// TIA Portal project "Semaforo Estruturado" (V16)

(* hardware
DEVICE "S7-1200 station_1"  S7-1200 Station
   slot 0: "Rack_0"  S7-1200 Rack  Rack  V1.0
   slot 1: "PLC_1"  CPU 1215C DC/DC/Rly  6ES7 215-1HG40-0XB0  V4.4
*)

// ===== PLC "PLC_1"  CPU 1215C DC/DC/Rly =====

VAR_GLOBAL   // PLC tag table "Default tag table"
   "Clock_Byte" AT %MB0 : Byte;
   "Clock_10Hz" AT %M0.0 : Bool;
   "Clock_5Hz" AT %M0.1 : Bool;
   "Clock_2.5Hz" AT %M0.2 : Bool;
   "Clock_2Hz" AT %M0.3 : Bool;
   "Clock_1.25Hz" AT %M0.4 : Bool;
   "Clock_1Hz" AT %M0.5 : Bool;
   "Clock_0.625Hz" AT %M0.6 : Bool;
   "Clock_0.5Hz" AT %M0.7 : Bool;
END_VAR

DATA_BLOCK "DB_Geral"   // DB1
{ S7_Optimized_Access := 'TRUE' }
VERSION : 0.1
   VAR
      Start : Bool;
      Stop : Bool;
      Reset : Bool;
      Estado : Bool;
      Time_of_Process : DInt;
      Time_PE_GroupA : Struct
         CutTimePE : DInt;
         TimePE : DInt := 20;
      END_STRUCT;
      Time_PE_GroupB : Struct
         CutTimePE : DInt;
         TimePE : DInt := 20;
      END_STRUCT;
      TimeOutCiclo : Struct
         "Estado 1" : DInt := 110;
         "Estado 2" : DInt := 120;
      END_STRUCT;
      ContadorGrupo : IEC_DCOUNTER;
   END_VAR
   VAR RETAIN
      PE : Struct
         GroupA : Bool;
         GroupB : Bool;
      END_STRUCT;
   END_VAR
   VAR
      Time_GroupA : Struct
         Red : Struct
            "begin" : DInt := 0;
            end : DInt := 40;
         END_STRUCT;
         Red_1 : Struct
            "begin" : DInt := 80;
            end : DInt := 110;
         END_STRUCT;
         Green : Struct
            "begin" : DInt := 40;
            end : DInt := 70;
         END_STRUCT;
         Yellow : Struct
            "begin" : DInt := 70;
            end : DInt := 80;
         END_STRUCT;
      END_STRUCT;
      Time_GroupB : Struct
         Red : Struct
            "begin" : DInt := 40;
            end : DInt := 110;
         END_STRUCT;
         Green : Struct
            "begin" : DInt := 0;
            end : DInt := 30;
         END_STRUCT;
         Yellow : Struct
            "begin" : DInt := 30;
            end : DInt := 40;
         END_STRUCT;
      END_STRUCT;
      Time_GroupC : Struct
         Red : Struct
            "begin" : DInt;
            end : DInt := 80;
         END_STRUCT;
         Green : Struct
            "begin" : DInt := 80;
            end : DInt := 100;
         END_STRUCT;
         Yellow : Struct
            "begin" : DInt := 100;
            end : DInt := 110;
         END_STRUCT;
      END_STRUCT;
   END_VAR
BEGIN
   ContadorGrupo.PV := 110;
END_DATA_BLOCK

DATA_BLOCK "DB_Input"   // DB2
{ S7_Optimized_Access := 'TRUE' }
VERSION : 0.1
   VAR
      Btn_PE_GroupA : Bool;
      Btn_PE_GroupB : Bool;
      Btn_Start : Bool;
      Btn_Stop : Bool;
      Btn_TestLamp : Bool;
      Btn_Reset : Bool;
   END_VAR
BEGIN
END_DATA_BLOCK

DATA_BLOCK "DB_Output"   // DB3
{ S7_Optimized_Access := 'TRUE' }
VERSION : 0.1
   VAR
      GroupA : Struct
         LampGreen : Bool;
         LampYell : Bool;
         LampRed : Bool;
      END_STRUCT;
      GroupB : Struct
         LampGreen : Bool;
         LampYell : Bool;
         LampRed : Bool;
      END_STRUCT;
      GroupC : Struct
         LampGreen : Bool;
         LampYell : Bool;
         LampRed : Bool;
      END_STRUCT;
      PE_GroupA : Struct
         LampGreen : Bool;
         LampRed : Bool;
      END_STRUCT;
      PE_GroupB : Struct
         LampGreen : Bool;
         LampRed : Bool;
      END_STRUCT;
   END_VAR
BEGIN
END_DATA_BLOCK

FUNCTION "FC_Geral" : Void   // FC1, LAD
{ S7_Optimized_Access := 'TRUE' }
VERSION : 0.1
   VAR_TEMP   // added for the SCL form of the ladder/FBD networks
      _w1 : Bool;
   END_VAR
BEGIN

REGION Network 1: Modo Start
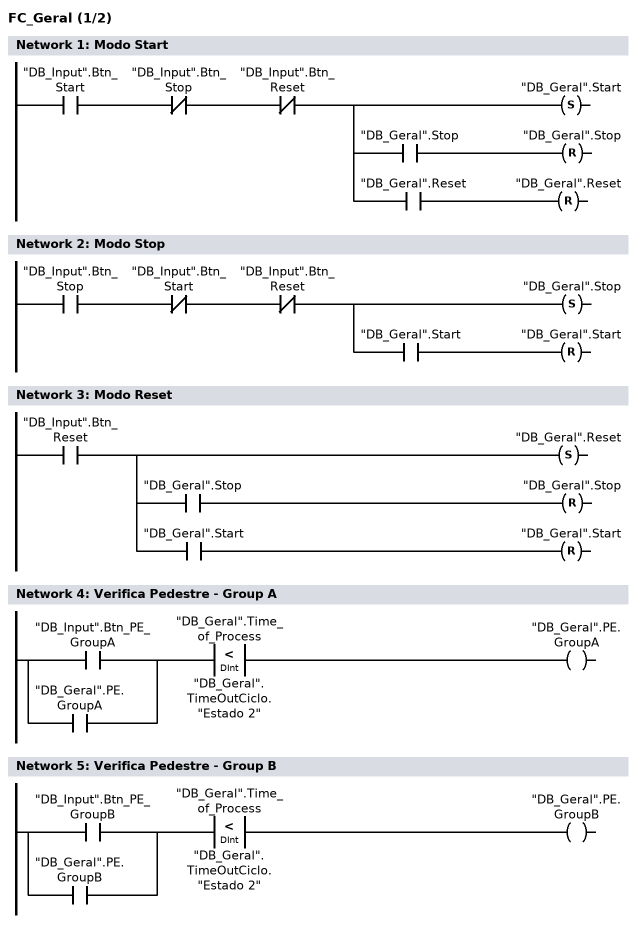
   RUNG wire#powerrail
      Contact( "DB_Input".Btn_Start )
      I_Contact( "DB_Input".Btn_Stop )
      I_Contact( "DB_Input".Btn_Reset )
      wire#w1
      S_Coil( "DB_Geral".Start )
   END_RUNG
   RUNG wire#w1
      Contact( "DB_Geral".Stop )
      R_Coil( "DB_Geral".Stop )
   END_RUNG
   RUNG wire#w1
      Contact( "DB_Geral".Reset )
      R_Coil( "DB_Geral".Reset )
   END_RUNG
   // the same network as SCL:
   #_w1 := "DB_Input".Btn_Start AND NOT "DB_Input".Btn_Stop AND NOT "DB_Input".Btn_Reset;
   IF #_w1 THEN "DB_Geral".Start := TRUE; END_IF;
   IF #_w1 AND "DB_Geral".Stop THEN "DB_Geral".Stop := FALSE; END_IF;
   IF #_w1 AND "DB_Geral".Reset THEN "DB_Geral".Reset := FALSE; END_IF;
END_REGION

REGION Network 2: Modo Stop
   RUNG wire#powerrail
      Contact( "DB_Input".Btn_Stop )
      I_Contact( "DB_Input".Btn_Start )
      I_Contact( "DB_Input".Btn_Reset )
      wire#w1
      S_Coil( "DB_Geral".Stop )
   END_RUNG
   RUNG wire#w1
      Contact( "DB_Geral".Start )
      R_Coil( "DB_Geral".Start )
   END_RUNG
   // the same network as SCL:
   #_w1 := "DB_Input".Btn_Stop AND NOT "DB_Input".Btn_Start AND NOT "DB_Input".Btn_Reset;
   IF #_w1 THEN "DB_Geral".Stop := TRUE; END_IF;
   IF #_w1 AND "DB_Geral".Start THEN "DB_Geral".Start := FALSE; END_IF;
END_REGION

REGION Network 3: Modo Reset
   RUNG wire#powerrail
      Contact( "DB_Input".Btn_Reset )
      wire#w1
      S_Coil( "DB_Geral".Reset )
   END_RUNG
   RUNG wire#w1
      Contact( "DB_Geral".Stop )
      R_Coil( "DB_Geral".Stop )
   END_RUNG
   RUNG wire#w1
      Contact( "DB_Geral".Start )
      R_Coil( "DB_Geral".Start )
   END_RUNG
   // the same network as SCL:
   IF "DB_Input".Btn_Reset THEN "DB_Geral".Reset := TRUE; END_IF;
   IF "DB_Input".Btn_Reset AND "DB_Geral".Stop THEN "DB_Geral".Stop := FALSE; END_IF;
   IF "DB_Input".Btn_Reset AND "DB_Geral".Start THEN "DB_Geral".Start := FALSE; END_IF;
END_REGION

REGION Network 4: Verifica Pedestre - Group A
   RUNG wire#powerrail
      Contact( "DB_Input".Btn_PE_GroupA )
      wire#w1
      { S7_Templates := "SrcType := DInt" } LT_Contact(in1 := "DB_Geral".Time_of_Process, in2 := "DB_Geral".TimeOutCiclo."Estado 2")
      Coil( "DB_Geral".PE.GroupA )
   END_RUNG
   RUNG wire#powerrail
      Contact( "DB_Geral".PE.GroupA )
   END_RUNG wire#w1
   // the same network as SCL:
   "DB_Geral".PE.GroupA := ("DB_Input".Btn_PE_GroupA OR "DB_Geral".PE.GroupA) AND ("DB_Geral".Time_of_Process < "DB_Geral".TimeOutCiclo."Estado 2");
END_REGION

REGION Network 5: Verifica Pedestre - Group B
   RUNG wire#powerrail
      Contact( "DB_Input".Btn_PE_GroupB )
      wire#w1
      { S7_Templates := "SrcType := DInt" } LT_Contact(in1 := "DB_Geral".Time_of_Process, in2 := "DB_Geral".TimeOutCiclo."Estado 2")
      Coil( "DB_Geral".PE.GroupB )
   END_RUNG
   RUNG wire#powerrail
      Contact( "DB_Geral".PE.GroupB )
   END_RUNG wire#w1
   // the same network as SCL:
   "DB_Geral".PE.GroupB := ("DB_Input".Btn_PE_GroupB OR "DB_Geral".PE.GroupB) AND ("DB_Geral".Time_of_Process < "DB_Geral".TimeOutCiclo."Estado 2");
END_REGION

REGION Network 6: Grupo A
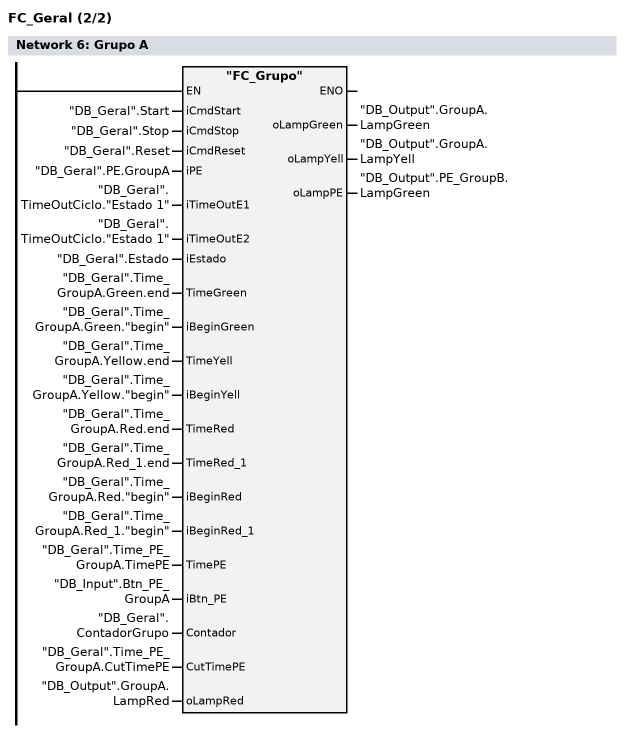
   RUNG wire#powerrail
      "FC_Grupo"(iCmdStart := "DB_Geral".Start, iCmdStop := "DB_Geral".Stop, iCmdReset := "DB_Geral".Reset, iPE := "DB_Geral".PE.GroupA, iTimeOutE1 := "DB_Geral".TimeOutCiclo."Estado 1", iTimeOutE2 := "DB_Geral".TimeOutCiclo."Estado 1", iEstado := "DB_Geral".Estado, TimeGreen := "DB_Geral".Time_GroupA.Green.end, iBeginGreen := "DB_Geral".Time_GroupA.Green."begin", TimeYell := "DB_Geral".Time_GroupA.Yellow.end, iBeginYell := "DB_Geral".Time_GroupA.Yellow."begin", TimeRed := "DB_Geral".Time_GroupA.Red.end, TimeRed_1 := "DB_Geral".Time_GroupA.Red_1.end, iBeginRed := "DB_Geral".Time_GroupA.Red."begin", iBeginRed_1 := "DB_Geral".Time_GroupA.Red_1."begin", TimePE := "DB_Geral".Time_PE_GroupA.TimePE, iBtn_PE := "DB_Input".Btn_PE_GroupA, Contador := "DB_Geral".ContadorGrupo, CutTimePE := "DB_Geral".Time_PE_GroupA.CutTimePE, oLampRed := "DB_Output".GroupA.LampRed, oLampGreen => "DB_Output".GroupA.LampGreen, oLampYell => "DB_Output".GroupA.LampYell, oLampPE => "DB_Output".PE_GroupB.LampGreen)
   END_RUNG
   // the same network as SCL:
   "FC_Grupo"(iCmdStart := "DB_Geral".Start,
              iCmdStop := "DB_Geral".Stop,
              iCmdReset := "DB_Geral".Reset,
              iPE := "DB_Geral".PE.GroupA,
              iTimeOutE1 := "DB_Geral".TimeOutCiclo."Estado 1",
              iTimeOutE2 := "DB_Geral".TimeOutCiclo."Estado 1",
              iEstado := "DB_Geral".Estado,
              TimeGreen := "DB_Geral".Time_GroupA.Green.end,
              iBeginGreen := "DB_Geral".Time_GroupA.Green."begin",
              TimeYell := "DB_Geral".Time_GroupA.Yellow.end,
              iBeginYell := "DB_Geral".Time_GroupA.Yellow."begin",
              TimeRed := "DB_Geral".Time_GroupA.Red.end,
              TimeRed_1 := "DB_Geral".Time_GroupA.Red_1.end,
              iBeginRed := "DB_Geral".Time_GroupA.Red."begin",
              iBeginRed_1 := "DB_Geral".Time_GroupA.Red_1."begin",
              TimePE := "DB_Geral".Time_PE_GroupA.TimePE,
              iBtn_PE := "DB_Input".Btn_PE_GroupA,
              Contador := "DB_Geral".ContadorGrupo,
              CutTimePE := "DB_Geral".Time_PE_GroupA.CutTimePE,
              oLampRed := "DB_Output".GroupA.LampRed,
              oLampGreen => "DB_Output".GroupA.LampGreen,
              oLampYell => "DB_Output".GroupA.LampYell,
              oLampPE => "DB_Output".PE_GroupB.LampGreen);
END_REGION
END_FUNCTION

FUNCTION "FC_Grupo" : Void   // FC2, LAD
{ S7_Optimized_Access := 'TRUE' }
VERSION : 0.1
   VAR_INPUT
      iCmdStart : Bool;
      iCmdStop : Bool;
      iCmdReset : Bool;
      iPE : Bool;
      iTimeOutE1 : DInt;
      iTimeOutE2 : DInt;
      iEstado : Bool;
      TimeGreen : DInt;
      iBeginGreen : DInt;
      TimeYell : DInt;
      iBeginYell : DInt;
      TimeRed : DInt;
      TimeRed_1 : DInt;
      iBeginRed : DInt;
      iBeginRed_1 : DInt;
      TimePE : DInt;
      iBtn_PE : Bool;
   END_VAR
   VAR_OUTPUT
      oLampGreen : Bool;
      oLampYell : Bool;
      oLampPE : Bool;
   END_VAR
   VAR_IN_OUT
      Contador : IEC_DCOUNTER;
      CutTimePE : DInt;
      oLampRed : Bool;
   END_VAR
BEGIN

REGION Network 1: Conta Tempo Fim de Ciclo
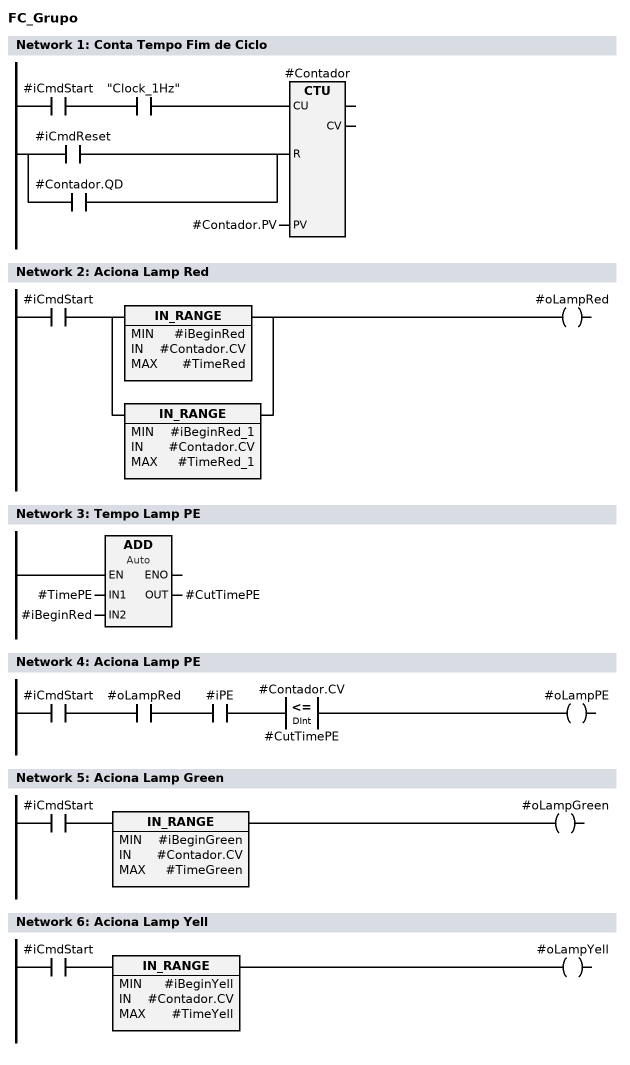
   #Contador.CTU(CU := #iCmdStart AND "Clock_1Hz", R := #iCmdReset OR #Contador.QD, PV := #Contador.PV);
END_REGION

REGION Network 2: Aciona Lamp Red
   RUNG wire#powerrail
      Contact( #iCmdStart )
      wire#w1
      { S7_Templates := "SrcType := DInt" } InRange(min := #iBeginRed, in := #Contador.CV, max := #TimeRed)
      wire#w2
      Coil( #oLampRed )
   END_RUNG
   RUNG wire#w1
      { S7_Templates := "SrcType := DInt" } InRange(min := #iBeginRed_1, in := #Contador.CV, max := #TimeRed_1)
   END_RUNG wire#w2
   // the same network as SCL:
   #oLampRed := #iCmdStart AND (((#iBeginRed <= #Contador.CV) AND (#Contador.CV <= #TimeRed)) OR ((#iBeginRed_1 <= #Contador.CV) AND (#Contador.CV <= #TimeRed_1)));
END_REGION

REGION Network 3: Tempo Lamp PE
   RUNG wire#powerrail
      Add(in1 := #TimePE, in2 := #iBeginRed, out => #CutTimePE)
   END_RUNG
   // the same network as SCL:
   #CutTimePE := #TimePE + #iBeginRed;
END_REGION

REGION Network 4: Aciona Lamp PE
   RUNG wire#powerrail
      Contact( #iCmdStart )
      Contact( #oLampRed )
      Contact( #iPE )
      { S7_Templates := "SrcType := DInt" } LE_Contact(in1 := #Contador.CV, in2 := #CutTimePE)
      Coil( #oLampPE )
   END_RUNG
   // the same network as SCL:
   #oLampPE := #iCmdStart AND #oLampRed AND #iPE AND (#Contador.CV <= #CutTimePE);
END_REGION

REGION Network 5: Aciona Lamp Green
   RUNG wire#powerrail
      Contact( #iCmdStart )
      { S7_Templates := "SrcType := DInt" } InRange(min := #iBeginGreen, in := #Contador.CV, max := #TimeGreen)
      Coil( #oLampGreen )
   END_RUNG
   // the same network as SCL:
   #oLampGreen := #iCmdStart AND (#iBeginGreen <= #Contador.CV) AND (#Contador.CV <= #TimeGreen);
END_REGION

REGION Network 6: Aciona Lamp Yell
   RUNG wire#powerrail
      Contact( #iCmdStart )
      { S7_Templates := "SrcType := DInt" } InRange(min := #iBeginYell, in := #Contador.CV, max := #TimeYell)
      Coil( #oLampYell )
   END_RUNG
   // the same network as SCL:
   #oLampYell := #iCmdStart AND (#iBeginYell <= #Contador.CV) AND (#Contador.CV <= #TimeYell);
END_REGION
END_FUNCTION

ORGANIZATION_BLOCK "Main"   // OB1, LAD, ProgramCycle
TITLE = "Main Program Sweep (Cycle)"
{ S7_Optimized_Access := 'TRUE' }
VERSION : 0.1
   VAR_INPUT
      Initial_Call : Bool;   // Initial call of this OB
      Remanence : Bool;   // =True, if remanent data are available
   END_VAR
BEGIN
END_ORGANIZATION_BLOCK